VERSION : 0.1
   VAR
      VFD_DELAY : Array[1..5] of IEC_TIMER;
   END_VAR
BEGIN
   VFD_DELAY[1].PT := T#10S;
   VFD_DELAY[2].PT := T#10S;
END_DATA_BLOCK

// folder: Timers/Totalizer/Datablocks

DATA_BLOCK "FT-1045_Totalizer_DB"   // DB7
{ S7_Optimized_Access := 'TRUE' }
VERSION : 0.1
// stored: InstanceOfName Totalizer_1
"Totalizer_1"
BEGIN
   interval := T#30s;
   cycle := T#500ms;
END_DATA_BLOCK

DATA_BLOCK "FT-1041_Totalizer_DB"   // DB88
{ S7_Optimized_Access := 'TRUE' }
VERSION : 0.1
// stored: InstanceOfName Totalizer_1
"Totalizer_1"
BEGIN
   cycle := T#500ms;
   interval := T#30s;
END_DATA_BLOCK

DATA_BLOCK "FT-2022_Totalizer_DB"   // DB111
{ S7_Optimized_Access := 'TRUE' }
VERSION : 0.1
// stored: InstanceOfName Totalizer_1
"Totalizer_1"
BEGIN
   cycle := T#500ms;
   interval := T#30s;
END_DATA_BLOCK

DATA_BLOCK "FT-2012_Totalizer_DB"   // DB112
{ S7_Optimized_Access := 'TRUE' }
VERSION : 0.1
// stored: InstanceOfName Totalizer_1
"Totalizer_1"
BEGIN
   interval := T#30s;
   cycle := T#500ms;
END_DATA_BLOCK

DATA_BLOCK "FT-2011_Totalizer_DB"   // DB113
{ S7_Optimized_Access := 'TRUE' }
VERSION : 0.1
// stored: InstanceOfName Totalizer_1
"Totalizer_1"
BEGIN
   interval := T#30s;
   cycle := T#500ms;
END_DATA_BLOCK

DATA_BLOCK "FT-1044_Totalizer_DB"   // DB114
{ S7_Optimized_Access := 'TRUE' }
VERSION : 0.1
// stored: InstanceOfName Totalizer_1
"Totalizer_1"
BEGIN
   interval := T#30s;
   cycle := T#500ms;
END_DATA_BLOCK

DATA_BLOCK "FT-1043_Totalizer_DB"   // DB115
{ S7_Optimized_Access := 'TRUE' }
VERSION : 0.1
// stored: InstanceOfName Totalizer_1
"Totalizer_1"
BEGIN
   interval := T#30s;
   cycle := T#500ms;
END_DATA_BLOCK

DATA_BLOCK "FT-1042_Totalizer_DB"   // DB116
{ S7_Optimized_Access := 'TRUE' }
VERSION : 0.1
// stored: InstanceOfName Totalizer_1
"Totalizer_1"
BEGIN
   interval := T#30s;
   cycle := T#500ms;
END_DATA_BLOCK

DATA_BLOCK "FT-3011_Totalizer_DB"   // DB117
{ S7_Optimized_Access := 'TRUE' }
VERSION : 0.1
// stored: InstanceOfName Totalizer_1
"Totalizer_1"
BEGIN
   interval := T#30s;
   cycle := T#500MS;
END_DATA_BLOCK

DATA_BLOCK "FT-2021_Totalizer_DB"   // DB118
{ S7_Optimized_Access := 'TRUE' }
VERSION : 0.1
// stored: InstanceOfName Totalizer_1
"Totalizer_1"
BEGIN
   interval := T#30s;
   cycle := T#500ms;
END_DATA_BLOCK

DATA_BLOCK "FT-1021_Totalizer_DB"   // DB190
{ S7_Optimized_Access := 'TRUE' }
VERSION : 0.1
// stored: InstanceOfName Totalizer_1
"Totalizer_1"
BEGIN
   interval := T#30s;
   cycle := T#500ms;
END_DATA_BLOCK

DATA_BLOCK "FT-1011_Totalizer_DB"   // DB254
{ S7_Optimized_Access := 'TRUE' }
VERSION : 0.1
// stored: InstanceOfName Totalizer_1
"Totalizer_1"
BEGIN
END_DATA_BLOCK

DATA_BLOCK "FT-3012_Totalizer_DB"   // DB376
{ S7_Optimized_Access := 'TRUE' }
VERSION : 0.1
// stored: InstanceOfName Totalizer_1
"Totalizer_1"
BEGIN
   interval := T#30s;
   cycle := T#500ms;
END_DATA_BLOCK

// folder: VFD/Datablocks

DATA_BLOCK "VFD-C301_DB"   // DB1
{ S7_Optimized_Access := 'TRUE' }
VERSION : 0.7
// stored: InstanceOfName VFD_Dumbdown
"VFD_Dumbdown"
BEGIN
END_DATA_BLOCK

DATA_BLOCK "VFD-C301R_DB"   // DB84
{ S7_Optimized_Access := 'TRUE' }
VERSION : 0.7
// stored: InstanceOfName VFD_Dumbdown
"VFD_Dumbdown"
BEGIN
END_DATA_BLOCK

DATA_BLOCK "VFD-R201_DB"   // DB85
{ S7_Optimized_Access := 'TRUE' }
VERSION : 0.7
// stored: InstanceOfName VFD_Dumbdown
"VFD_Dumbdown"
BEGIN
   Motor_max_RPM := 450.0;
END_DATA_BLOCK

DATA_BLOCK "VFD-T103_DB"   // DB107
{ S7_Optimized_Access := 'TRUE' }
VERSION : 0.7
// stored: InstanceOfName VFD_Dumbdown
"VFD_Dumbdown"
BEGIN
END_DATA_BLOCK

DATA_BLOCK "VFD-T102A_DB"   // DB108
{ S7_Optimized_Access := 'TRUE' }
VERSION : 0.7
// stored: InstanceOfName VFD_Dumbdown
"VFD_Dumbdown"
BEGIN
   Motor_max_RPM := 1770.0;
END_DATA_BLOCK

DATA_BLOCK "VFD-T101A_DB"   // DB109
{ S7_Optimized_Access := 'TRUE' }
VERSION : 0.7
// stored: InstanceOfName VFD_Dumbdown
"VFD_Dumbdown"
BEGIN
   Motor_max_RPM := 1730.0;
END_DATA_BLOCK

DATA_BLOCK "VFD-R202_DB"   // DB110
{ S7_Optimized_Access := 'TRUE' }
VERSION : 0.7
// stored: InstanceOfName VFD_Dumbdown
"VFD_Dumbdown"
BEGIN
   Motor_max_RPM := 450.0;
END_DATA_BLOCK

DATA_BLOCK "VFD-T101B_DB"   // DB183
{ S7_Optimized_Access := 'TRUE' }
VERSION : 0.7
// stored: InstanceOfName VFD_Dumbdown
"VFD_Dumbdown"
BEGIN
   Motor_max_RPM := 1730.0;
END_DATA_BLOCK

DATA_BLOCK "VFD-T102B_DB"   // DB184
{ S7_Optimized_Access := 'TRUE' }
VERSION : 0.7
// stored: InstanceOfName VFD_Dumbdown
"VFD_Dumbdown"
BEGIN
   Motor_max_RPM := 1770.0;
END_DATA_BLOCK

// folder: VFD/T103_VFD

DATA_BLOCK "T103_VFD_Control_DB"   // DB263
{ S7_Optimized_Access := 'TRUE' }
VERSION : 0.1
   VAR
      AutoSpeedSP : Real;   // Auto Speed SP
   END_VAR
BEGIN
END_DATA_BLOCK

DATA_BLOCK "VFD_T103_PN_DB"   // DB264
{ S7_Optimized_Access := 'TRUE' }
VERSION : 0.1
// stored: InstanceOfName VFD_PNCtrl
"VFD_PNCtrl"
BEGIN
END_DATA_BLOCK

// folder: Valves/Control Valves

DATA_BLOCK "FV-4012_DB"   // DB177
{ S7_Optimized_Access := 'TRUE' }
VERSION : 0.1
// stored: InstanceOfName Valve-CV
"Valve-CV"
BEGIN
END_DATA_BLOCK

// folder: Valves/Control Valves/Datablocks

DATA_BLOCK "FV-2011_DB"   // DB80
{ S7_Optimized_Access := 'TRUE' }
VERSION : 0.1
// stored: InstanceOfName Valve-CV
"Valve-CV"
BEGIN
END_DATA_BLOCK

DATA_BLOCK "FV-2012_DB"   // DB81
{ S7_Optimized_Access := 'TRUE' }
VERSION : 0.1
// stored: InstanceOfName Valve-CV
"Valve-CV"
BEGIN
END_DATA_BLOCK

DATA_BLOCK "FV-2021_DB"   // DB82
{ S7_Optimized_Access := 'TRUE' }
VERSION : 0.1
// stored: InstanceOfName Valve-CV
"Valve-CV"
BEGIN
END_DATA_BLOCK

DATA_BLOCK "FV-2022_DB"   // DB83
{ S7_Optimized_Access := 'TRUE' }
VERSION : 0.1
// stored: InstanceOfName Valve-CV
"Valve-CV"
BEGIN
END_DATA_BLOCK

DATA_BLOCK "FV-3011_DB"   // DB234
{ S7_Optimized_Access := 'TRUE' }
VERSION : 0.1
// stored: InstanceOfName Valve-CV
"Valve-CV"
BEGIN
END_DATA_BLOCK

DATA_BLOCK "FV-4011_DB"   // DB381
{ S7_Optimized_Access := 'TRUE' }
VERSION : 0.1
// stored: InstanceOfName Valve-CV
"Valve-CV"
BEGIN
END_DATA_BLOCK

DATA_BLOCK "FV-4021_DB"   // DB418
{ S7_Optimized_Access := 'TRUE' }
VERSION : 0.1
// stored: InstanceOfName Valve-CV
"Valve-CV"
BEGIN
END_DATA_BLOCK

DATA_BLOCK "FV-4024_DB"   // DB419
{ S7_Optimized_Access := 'TRUE' }
VERSION : 0.1
// stored: InstanceOfName Valve-CV
"Valve-CV"
BEGIN
END_DATA_BLOCK

DATA_BLOCK "FV-4025_DB"   // DB420
{ S7_Optimized_Access := 'TRUE' }
VERSION : 0.1
// stored: InstanceOfName Valve-CV
"Valve-CV"
BEGIN
END_DATA_BLOCK

// folder: Valves/Solenoid Valve/Datablocks

DATA_BLOCK "XV-1033_DB"   // DB2
{ S7_Optimized_Access := 'FALSE' }
VERSION : 1.0
// stored: InstanceOfName Valve-SV
"Valve-SV"
BEGIN
   EM := 1;
END_DATA_BLOCK

DATA_BLOCK "XV-1041_DB"   // DB3
{ S7_Optimized_Access := 'FALSE' }
VERSION : 1.0
// stored: InstanceOfName Valve-SV
"Valve-SV"
BEGIN
   EM := 1;
END_DATA_BLOCK

DATA_BLOCK "XV-1011_DB"   // DB4
{ S7_Optimized_Access := 'FALSE' }
VERSION : 1.0
// stored: InstanceOfName Valve-SV
"Valve-SV"
BEGIN
   EM := 1;
END_DATA_BLOCK

DATA_BLOCK "XV-1013_DB"   // DB5
{ S7_Optimized_Access := 'FALSE' }
VERSION : 1.0
// stored: InstanceOfName Valve-SV
"Valve-SV"
BEGIN
   EM := 1;
END_DATA_BLOCK

DATA_BLOCK "XV-1021_DB"   // DB10
{ S7_Optimized_Access := 'FALSE' }
VERSION : 1.0
// stored: InstanceOfName Valve-SV
"Valve-SV"
BEGIN
   EM := 1;
END_DATA_BLOCK

DATA_BLOCK "XV-1043_DB"   // DB12
{ S7_Optimized_Access := 'FALSE' }
VERSION : 1.0
// stored: InstanceOfName Valve-SV
"Valve-SV"
BEGIN
   EM := 1;
END_DATA_BLOCK

DATA_BLOCK "XV-1044_DB"   // DB13
{ S7_Optimized_Access := 'FALSE' }
VERSION : 1.0
// stored: InstanceOfName Valve-SV
"Valve-SV"
BEGIN
   EM := 1;
END_DATA_BLOCK

DATA_BLOCK "XV-2011_DB"   // DB14
{ S7_Optimized_Access := 'FALSE' }
VERSION : 1.0
// stored: InstanceOfName Valve-SV
"Valve-SV"
BEGIN
   EM := 1;
END_DATA_BLOCK

DATA_BLOCK "XV-2012_DB"   // DB15
{ S7_Optimized_Access := 'FALSE' }
VERSION : 1.0
// stored: InstanceOfName Valve-SV
"Valve-SV"
BEGIN
   EM := 1;
END_DATA_BLOCK

DATA_BLOCK "XV-2013_DB"   // DB16
{ S7_Optimized_Access := 'FALSE' }
VERSION : 1.0
// stored: InstanceOfName Valve-SV
"Valve-SV"
BEGIN
   EM := 1;
END_DATA_BLOCK

DATA_BLOCK "XV-2021_DB"   // DB18
{ S7_Optimized_Access := 'FALSE' }
VERSION : 1.0
// stored: InstanceOfName Valve-SV
"Valve-SV"
BEGIN
   EM := 1;
END_DATA_BLOCK

DATA_BLOCK "XV-2023_DB"   // DB19
{ S7_Optimized_Access := 'FALSE' }
VERSION : 1.0
// stored: InstanceOfName Valve-SV
"Valve-SV"
BEGIN
   EM := 1;
END_DATA_BLOCK

DATA_BLOCK "XV-1032_DB"   // DB21
{ S7_Optimized_Access := 'FALSE' }
VERSION : 1.0
// stored: InstanceOfName Valve-SV
"Valve-SV"
BEGIN
   EM := 1;
END_DATA_BLOCK

DATA_BLOCK "XV-3011_DB"   // DB22
{ S7_Optimized_Access := 'FALSE' }
VERSION : 1.0
// stored: InstanceOfName Valve-SV
"Valve-SV"
BEGIN
   EM := 1;
END_DATA_BLOCK

DATA_BLOCK "XV-3012_DB"   // DB23
{ S7_Optimized_Access := 'FALSE' }
VERSION : 1.0
// stored: InstanceOfName Valve-SV
"Valve-SV"
BEGIN
   EM := 1;
END_DATA_BLOCK

DATA_BLOCK "XV-3013_DB"   // DB24
{ S7_Optimized_Access := 'FALSE' }
VERSION : 1.0
// stored: InstanceOfName Valve-SV
"Valve-SV"
BEGIN
   EM := 1;
END_DATA_BLOCK

DATA_BLOCK "XV-1045_DB"   // DB25
{ S7_Optimized_Access := 'FALSE' }
VERSION : 1.0
// stored: InstanceOfName Valve-SV
"Valve-SV"
BEGIN
   EM := 1;
END_DATA_BLOCK

DATA_BLOCK "XV-1023_DB"   // DB27
{ S7_Optimized_Access := 'FALSE' }
VERSION : 1.0
// stored: InstanceOfName Valve-SV
"Valve-SV"
BEGIN
   EM := 1;
END_DATA_BLOCK

DATA_BLOCK "XV-4024_DB"   // DB28
{ S7_Optimized_Access := 'FALSE' }
VERSION : 1.0
// stored: InstanceOfName Valve-SV
"Valve-SV"
BEGIN
   EM := 1;
END_DATA_BLOCK

DATA_BLOCK "XV-4025_DB"   // DB29
{ S7_Optimized_Access := 'FALSE' }
VERSION : 1.0
// stored: InstanceOfName Valve-SV
"Valve-SV"
BEGIN
   EM := 1;
END_DATA_BLOCK

DATA_BLOCK "XV-1042_DB"   // DB99
{ S7_Optimized_Access := 'FALSE' }
VERSION : 1.0
// stored: InstanceOfName Valve-SV
"Valve-SV"
BEGIN
   EM := 1;
END_DATA_BLOCK

DATA_BLOCK "XV-2022_DB"   // DB104
{ S7_Optimized_Access := 'FALSE' }
VERSION : 1.0
// stored: InstanceOfName Valve-SV
"Valve-SV"
BEGIN
   EM := 1;
END_DATA_BLOCK

DATA_BLOCK "XV-1031_DB"   // DB106
{ S7_Optimized_Access := 'FALSE' }
VERSION : 1.0
// stored: InstanceOfName Valve-SV
"Valve-SV"
BEGIN
   EM := 1;
END_DATA_BLOCK

DATA_BLOCK "XV-4021_DB"   // DB416
{ S7_Optimized_Access := 'FALSE' }
VERSION : 1.0
// stored: InstanceOfName Valve-SV
"Valve-SV"
BEGIN
END_DATA_BLOCK

DATA_BLOCK "XV-4022_DB"   // DB417
{ S7_Optimized_Access := 'FALSE' }
VERSION : 1.0
// stored: InstanceOfName Valve-SV
"Valve-SV"
BEGIN
END_DATA_BLOCK

// folder: 0)Organization Blocks

ORGANIZATION_BLOCK "Main"   // OB1, LAD, ProgramCycle
TITLE = "Main Program Sweep (Cycle)"
{ S7_Optimized_Access := 'TRUE' }
VERSION : 0.1
// Updated Date:
// Note:
   VAR_INPUT
      Initial_Call : Bool;   // Initial call of this OB
      Remanence : Bool;   // =True, if remanent data are available
   END_VAR
   VAR_TEMP
      "bool" : Bool;
   END_VAR
   VAR CONSTANT
      Idle_Star : Int := 0;
      Idle_End : Int := 49;
      Shutdown_Star : Int := 50;
      Shutdown_End : Int := 99;
      Inititilize_Start : Int := 100;
      Inititilize_End : Int := 199;
   END_VAR
BEGIN

REGION Network 1: Interlocks & Diagnostic
   // Interlocks_FC: Contains all interlock Sequences 
   // Diag_FC: Contains all diagnostic  Sequences
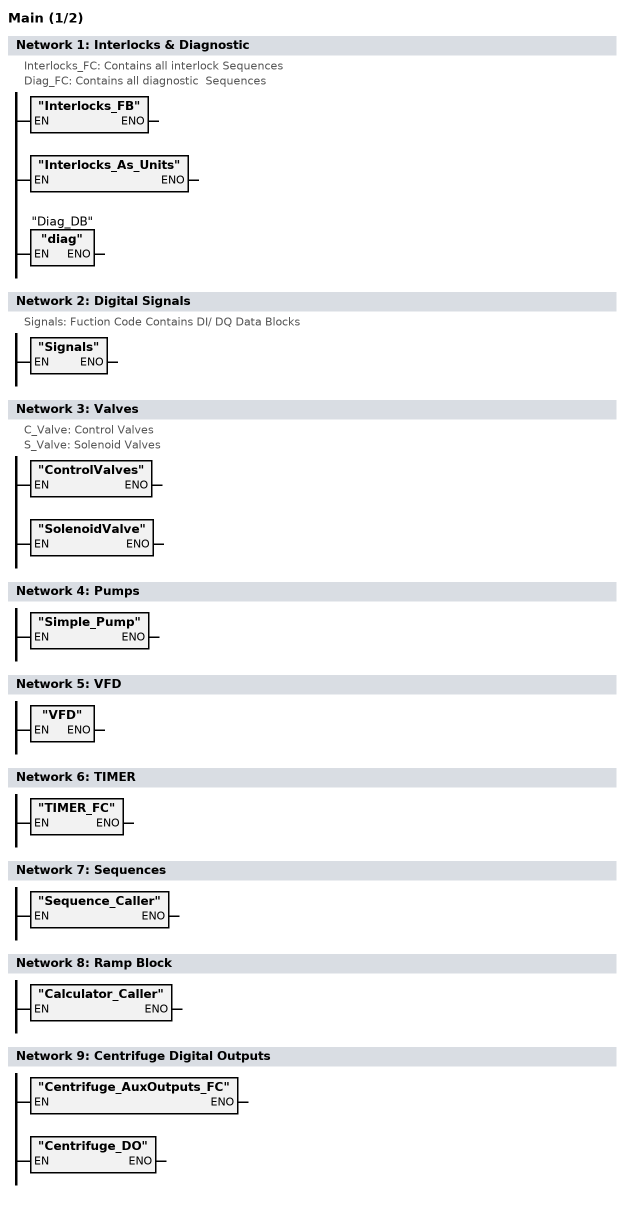
   RUNG wire#powerrail
      "Interlocks_FB"()
   END_RUNG
   RUNG wire#powerrail
      "Interlocks_As_Units"()
   END_RUNG
   RUNG wire#powerrail
      "Diag_DB"()
   END_RUNG
   // the same network as SCL:
   "Interlocks_FB"();
   "Interlocks_As_Units"();
   "Diag_DB"();   // "diag"
END_REGION

REGION Network 2: Digital Signals
   // Signals: Fuction Code Contains DI/ DQ Data Blocks
   RUNG wire#powerrail
      "Signals"()
   END_RUNG
   // the same network as SCL:
   "Signals"();
END_REGION

REGION Network 3: Valves
   // C_Valve: Control Valves 
   // S_Valve: Solenoid Valves
   RUNG wire#powerrail
      "ControlValves"()
   END_RUNG
   RUNG wire#powerrail
      "SolenoidValve"()
   END_RUNG
   // the same network as SCL:
   "ControlValves"();
   "SolenoidValve"();
END_REGION

REGION Network 4: Pumps
   RUNG wire#powerrail
      "Simple_Pump"()
   END_RUNG
   // the same network as SCL:
   "Simple_Pump"();
END_REGION

REGION Network 5: VFD
   RUNG wire#powerrail
      "VFD"()
   END_RUNG
   // the same network as SCL:
   "VFD"();
END_REGION

REGION Network 6: TIMER
   RUNG wire#powerrail
      "TIMER_FC"()
   END_RUNG
   // the same network as SCL:
   "TIMER_FC"();
END_REGION

REGION Network 7: Sequences
   RUNG wire#powerrail
      "Sequence_Caller"()
   END_RUNG
   // the same network as SCL:
   "Sequence_Caller"();
END_REGION

REGION Network 8: Ramp Block
   RUNG wire#powerrail
      "Calculator_Caller"()
   END_RUNG
   // the same network as SCL:
   "Calculator_Caller"();
END_REGION

REGION Network 9: Centrifuge Digital Outputs
   RUNG wire#powerrail
      "Centrifuge_AuxOutputs_FC"()
   END_RUNG
   RUNG wire#powerrail
      "Centrifuge_DO"()
   END_RUNG
   // the same network as SCL:
   "Centrifuge_AuxOutputs_FC"();
   "Centrifuge_DO"();
END_REGION

REGION Network 10: Cause and Effect Matrix
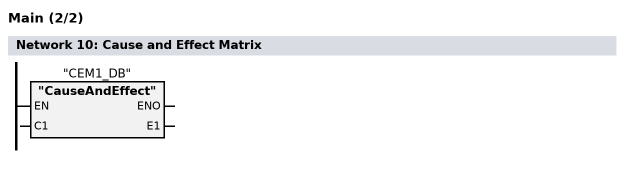
   RUNG wire#powerrail
      "CEM1_DB"(C1 :=, E1 =>)
   END_RUNG
   // the same network as SCL:
   "CEM1_DB"();   // "CauseAndEffect"
END_REGION
END_ORGANIZATION_BLOCK

ORGANIZATION_BLOCK "Cycle_5s"   // OB30, LAD, CyclicInterrupt
{ S7_Optimized_Access := 'TRUE' }
VERSION : 0.1
   VAR_INPUT
      Initial_Call : Bool;   // Initial call of this OB
      Event_Count : Int;   // Events discarded
   END_VAR
BEGIN

REGION Network 1: Temperature Trasmitters
   // Temperature Trasmitters Function Code
END_REGION
END_ORGANIZATION_BLOCK

ORGANIZATION_BLOCK "Cycle_100ms"   // OB31, LAD, CyclicInterrupt
{ S7_Optimized_Access := 'TRUE' }
VERSION : 0.1
   VAR_INPUT
      Initial_Call : Bool;   // Initial call of this OB
      Event_Count : Int;   // Events discarded
   END_VAR
   VAR_TEMP   // added for the SCL form of the ladder/FBD networks
      _w1 : Bool;
      _w2 : Bool;
      _w3 : Bool;
   END_VAR
BEGIN

REGION Network 1: PH Trasmitters
   // PH Trasmitters Function Code
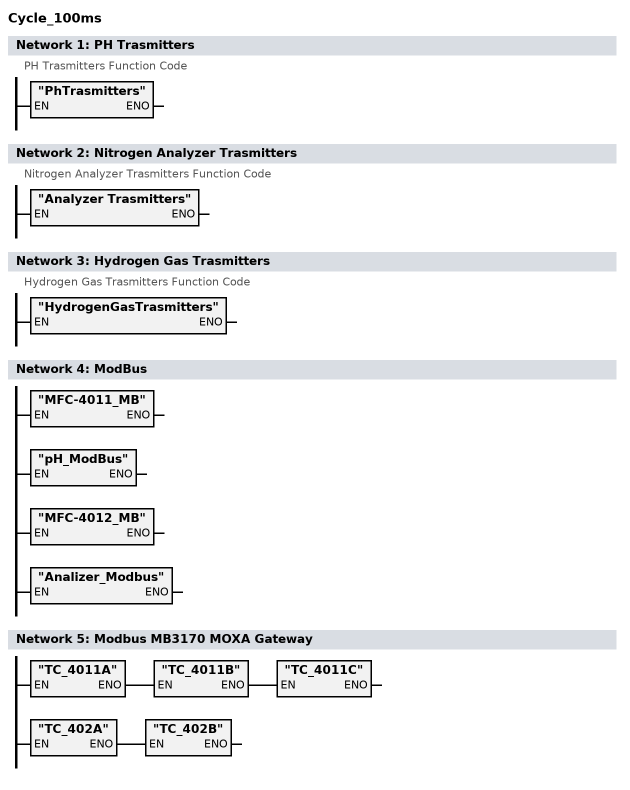
   RUNG wire#powerrail
      "PhTrasmitters"()
   END_RUNG
   // the same network as SCL:
   "PhTrasmitters"();
END_REGION

REGION Network 2: Nitrogen Analyzer Trasmitters
   // Nitrogen Analyzer Trasmitters Function Code
   RUNG wire#powerrail
      "Analyzer Trasmitters"()
   END_RUNG
   // the same network as SCL:
   "Analyzer Trasmitters"();
END_REGION

REGION Network 3: Hydrogen Gas Trasmitters
   // Hydrogen Gas Trasmitters Function Code
   RUNG wire#powerrail
      "HydrogenGasTrasmitters"()
   END_RUNG
   // the same network as SCL:
   "HydrogenGasTrasmitters"();
END_REGION

REGION Network 4: ModBus
   RUNG wire#powerrail
      "MFC-4011_MB"()
   END_RUNG
   RUNG wire#powerrail
      "pH_ModBus"()
   END_RUNG
   RUNG wire#powerrail
      "MFC-4012_MB"()
   END_RUNG
   RUNG wire#powerrail
      "Analizer_Modbus"()
   END_RUNG
   // the same network as SCL:
   "MFC-4011_MB"();
   "pH_ModBus"();
   "MFC-4012_MB"();
   "Analizer_Modbus"();
END_REGION

REGION Network 5: Modbus MB3170 MOXA Gateway
   RUNG wire#powerrail
      "TC_4011A"()
      "TC_4011B"()
      "TC_4011C"()
   END_RUNG
   RUNG wire#powerrail
      "TC_402A"()
      "TC_402B"()
   END_RUNG
   // the same network as SCL:
   "TC_4011A"(ENO => #_w1);
   "TC_4011B"(EN := #_w1, ENO => #_w2);
   IF #_w2 THEN "TC_4011C"(); END_IF;
   "TC_402A"(ENO => #_w3);
   IF #_w3 THEN "TC_402B"(); END_IF;
END_REGION
END_ORGANIZATION_BLOCK

ORGANIZATION_BLOCK "Cycle_1s"   // OB32, LAD, CyclicInterrupt
TITLE = Cyclic interrupt (Cycle) 1 Second"
{ S7_Optimized_Access := 'TRUE' }
VERSION : 0.1
   VAR_INPUT
      Initial_Call : Bool;   // Initial call of this OB
      Event_Count : Int;   // Events discarded
   END_VAR
BEGIN

REGION Network 1: PIDController
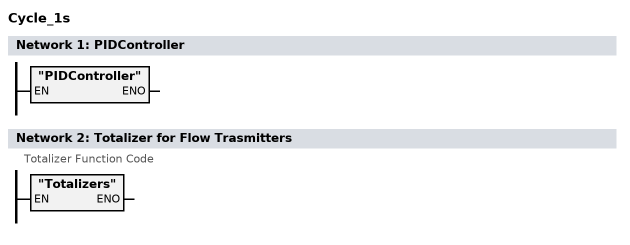
   RUNG wire#powerrail
      "PIDController"()
   END_RUNG
   // the same network as SCL:
   "PIDController"();
END_REGION

REGION Network 2: Totalizer for Flow Trasmitters
   // Totalizer Function Code
   RUNG wire#powerrail
      "Totalizers"()
   END_RUNG
   // the same network as SCL:
   "Totalizers"();
END_REGION
END_ORGANIZATION_BLOCK

ORGANIZATION_BLOCK "Cycle_500ms"   // OB33, LAD, CyclicInterrupt
{ S7_Optimized_Access := 'TRUE' }
VERSION : 0.1
   VAR_INPUT
      Initial_Call : Bool;   // Initial call of this OB
      Event_Count : Int;   // Events discarded
   END_VAR
   VAR_TEMP
      "REAL_R-201" : Real;
      "INT_R-201" : Real;
      "INT_R-202" : Real;
      "REAL_R-202" : Real;
   END_VAR
BEGIN

REGION Network 1: Flow Trasmitters
   // Flow Trasmitters Function Code
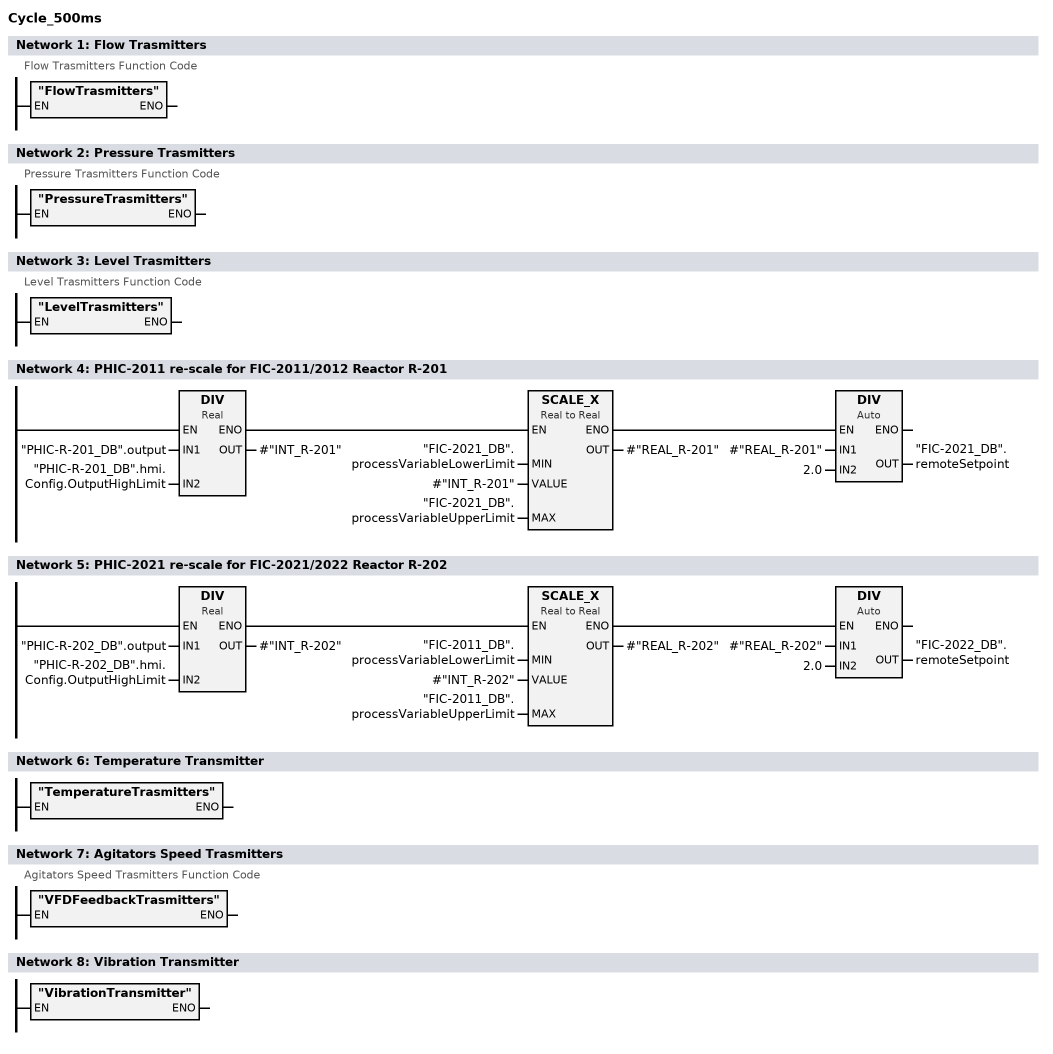
   RUNG wire#powerrail
      "FlowTrasmitters"()
   END_RUNG
   // the same network as SCL:
   "FlowTrasmitters"();
END_REGION

REGION Network 2: Pressure Trasmitters
   // Pressure Trasmitters Function Code
   RUNG wire#powerrail
      "PressureTrasmitters"()
   END_RUNG
   // the same network as SCL:
   "PressureTrasmitters"();
END_REGION

REGION Network 3: Level Trasmitters
   // Level Trasmitters Function Code
   RUNG wire#powerrail
      "LevelTrasmitters"()
   END_RUNG
   // the same network as SCL:
   "LevelTrasmitters"();
END_REGION

REGION Network 4: PHIC-2011 re-scale for FIC-2011/2012 Reactor R-201
   RUNG wire#powerrail
      { S7_Templates := "SrcType := Real"; S7_GenerateENO := "TRUE" } Div(in1 := "PHIC-R-201_DB".output, in2 := "PHIC-R-201_DB".hmi.Config.OutputHighLimit, out => #"INT_R-201")
      { S7_Templates := "[SrcType := Real, DestType := Real]"; S7_GenerateENO := "TRUE" } Scale(min := "FIC-2021_DB".processVariableLowerLimit, value := #"INT_R-201", max := "FIC-2021_DB".processVariableUpperLimit, out => #"REAL_R-201")
      { S7_GenerateENO := "TRUE" } Div(in1 := #"REAL_R-201", in2 := 2.0, out => "FIC-2021_DB".remoteSetpoint)
   END_RUNG
   // the same network as SCL:
   // ENO of a box is taken as its EN; it also drops when the box reports an error
   #"INT_R-201" := "PHIC-R-201_DB".output / "PHIC-R-201_DB".hmi.Config.OutputHighLimit;
   #"REAL_R-201" := SCALE_X(MIN := "FIC-2021_DB".processVariableLowerLimit, VALUE := #"INT_R-201", MAX := "FIC-2021_DB".processVariableUpperLimit);
   "FIC-2021_DB".remoteSetpoint := #"REAL_R-201" / 2.0;
END_REGION

REGION Network 5: PHIC-2021 re-scale for FIC-2021/2022 Reactor R-202
   RUNG wire#powerrail
      { S7_Templates := "SrcType := Real"; S7_GenerateENO := "TRUE" } Div(in1 := "PHIC-R-202_DB".output, in2 := "PHIC-R-202_DB".hmi.Config.OutputHighLimit, out => #"INT_R-202")
      { S7_Templates := "[SrcType := Real, DestType := Real]"; S7_GenerateENO := "TRUE" } Scale(min := "FIC-2011_DB".processVariableLowerLimit, value := #"INT_R-202", max := "FIC-2011_DB".processVariableUpperLimit, out => #"REAL_R-202")
      { S7_GenerateENO := "TRUE" } Div(in1 := #"REAL_R-202", in2 := 2.0, out => "FIC-2022_DB".remoteSetpoint)
   END_RUNG
   // the same network as SCL:
   // ENO of a box is taken as its EN; it also drops when the box reports an error
   #"INT_R-202" := "PHIC-R-202_DB".output / "PHIC-R-202_DB".hmi.Config.OutputHighLimit;
   #"REAL_R-202" := SCALE_X(MIN := "FIC-2011_DB".processVariableLowerLimit, VALUE := #"INT_R-202", MAX := "FIC-2011_DB".processVariableUpperLimit);
   "FIC-2022_DB".remoteSetpoint := #"REAL_R-202" / 2.0;
END_REGION

REGION Network 6: Temperature Transmitter
   RUNG wire#powerrail
      "TemperatureTrasmitters"()
   END_RUNG
   // the same network as SCL:
   "TemperatureTrasmitters"();
END_REGION

REGION Network 7: Agitators Speed Trasmitters
   // Agitators Speed Trasmitters Function Code
   RUNG wire#powerrail
      "VFDFeedbackTrasmitters"()
   END_RUNG
   // the same network as SCL:
   "VFDFeedbackTrasmitters"();
END_REGION

REGION Network 8: Vibration Transmitter
   RUNG wire#powerrail
      "VibrationTransmitter"()
   END_RUNG
   // the same network as SCL:
   "VibrationTransmitter"();
END_REGION
END_ORGANIZATION_BLOCK

ORGANIZATION_BLOCK "CPU redundancy error"   // OB72, LAD, CPURedundancyError
{ S7_Optimized_Access := 'TRUE' }
VERSION : 0.1
   VAR_INPUT
      LADDR : Hw_Any;   // Hardware identifier of the local device
      Event_Class : Byte;   // according to S7 classic
      Fault_ID : Byte;   // Fault_ID as in S7 classic
   END_VAR
BEGIN
END_ORGANIZATION_BLOCK

ORGANIZATION_BLOCK "Diagnostic error interrupt"   // OB82, LAD, DiagnosticErrorInterrupt
{ S7_Optimized_Access := 'TRUE' }
VERSION : 0.1
   VAR_INPUT
      IO_State : Word;   // IO state of the HW object
      LADDR : Hw_Any;   // Hardware identifier
      Channel : UInt;   // Channel number
      MultiError : Bool;   // =true if more than one error is present
   END_VAR
BEGIN
END_ORGANIZATION_BLOCK

ORGANIZATION_BLOCK "Startup"   // OB100, LAD, Startup
TITLE = "Complete Restart"
{ S7_Optimized_Access := 'TRUE' }
VERSION : 0.1
   VAR_INPUT
      LostRetentive : Bool;   // True if retentive data are lost
      LostRTC : Bool;   // True if date and time are lost
   END_VAR
BEGIN

REGION Network 1: VFD Set to Automode
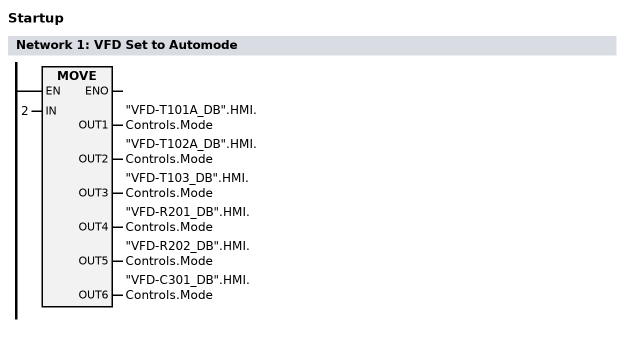
   RUNG wire#powerrail
      { S7_GenerateENO := "TRUE" } Move(in := 2, out1 => "VFD-T101A_DB".HMI.Controls.Mode, out2 => "VFD-T102A_DB".HMI.Controls.Mode, out3 => "VFD-T103_DB".HMI.Controls.Mode, out4 => "VFD-R201_DB".HMI.Controls.Mode, out5 => "VFD-R202_DB".HMI.Controls.Mode, out6 => "VFD-C301_DB".HMI.Controls.Mode)
   END_RUNG
   // the same network as SCL:
   "VFD-T101A_DB".HMI.Controls.Mode := 2;
   "VFD-T102A_DB".HMI.Controls.Mode := 2;
   "VFD-T103_DB".HMI.Controls.Mode := 2;
   "VFD-R201_DB".HMI.Controls.Mode := 2;
   "VFD-R202_DB".HMI.Controls.Mode := 2;
   "VFD-C301_DB".HMI.Controls.Mode := 2;
END_REGION
END_ORGANIZATION_BLOCK

ORGANIZATION_BLOCK "Programming error"   // OB121, LAD, ProgrammingError
{ S7_Optimized_Access := 'TRUE' }
VERSION : 0.1
   VAR_INPUT
      BlockNr : UInt;   // Number of causing block
      Reaction : USInt;   // 0:ignore, 1:substitute, 2:skip
      Fault_ID : Byte;   // Fault identifier
      BlockType : USInt;   // 16#01:OB, 16#02:FC, 16#03:FB, 16#04:SFC, 16#05:SFB, 16#06:DB: Type of block causing the error
      Area : USInt;   // Area where the error occured
      DBNr : DB_ANY;   // DB number if Area = DB or DI
      Csg_OBNr : OB_Any;   // Number of OB causing the error
      Csg_Prio : USInt;   // Priority of OB causing the error
      Width : USInt;   // 0:bit, 1:byte, 2:word, 3:dword, 4:lword
   END_VAR
BEGIN
END_ORGANIZATION_BLOCK

ORGANIZATION_BLOCK "IO access error"   // OB122, LAD, IOAccessError
{ S7_Optimized_Access := 'TRUE' }
VERSION : 0.1
   VAR_INPUT
      BlockNr : UInt;   // Number of causing block
      Reaction : USInt;   // 0:ignore, 1:substitute, 2:skip
      Fault_ID : Byte;   // 16#42:reading, 16#43:writing
      BlockType : USInt;   // 16#01:OB, 16#02:FC, 16#03:FB, 16#04:SFC, 16#05:SFB, 16#06:DB: Type of block causing the error
      Area : USInt;   // 16#81:I, 16#82:Q: IO area where the IOaccess error occured
      DBNr : DB_ANY;   // Reserved for system
      Csg_OBNr : OB_Any;   // Number of OB causing the error
      Csg_Prio : USInt;   // Priority of OB causing the error
      Width : USInt;   // 0:bit, 1:byte, 2:word, 3:dword, 4:lword
   END_VAR
BEGIN
END_ORGANIZATION_BLOCK

// folder: 1}Library

FUNCTION_BLOCK "UPS1600"   // FB15, LAD
{ S7_Optimized_Access := 'TRUE' }
VERSION : 0.1
   VAR_INPUT
      addrIn : Hw_Io := 260;   // HW-address of the UPS1600 must be insert there
      cyclicIOAddr : Hw_Io;   // IO Data submodule address must be inserted here
      upsExecuteReset : Bool;   // Input must be set if the station is ready for shutdown <- the station/ partners are ready to deactivate the tension
   END_VAR
   VAR_OUTPUT
      upsReadyForReset : Bool := False;   // Output will be set if the Block timer elapse -> signal to shutdown the station/ partners
   END_VAR
   VAR
      HMI : Struct
         Mode : Struct
            bufferMode : Byte := 16#80;   // Buffer mode //Value range: 0 = active, 255 = inactive
            readyForBuffering : Byte;   // Buffer readiness //Value range: 0=FALSE, 255=TRUE
         END_STRUCT;
         State : Struct
            Details : Struct
               orderNumber : String[20];   // Article no.
               serialNumber : String[20];   // Serial number
               deviceName : String[20];   // Name of the device
               versionNumber : String[30];   // Version number
               deviceHwRevision : Int;   // HW revision
               deviceSwRevision1 : Byte;   // SW revision1
               deviceSwRevision2 : Byte;   // SW revision2
               deviceSwRevision3 : Byte;   // Sw revision3
               batFamily : Byte;   // Battery family //Value range: BAT1600 = 1, UPS1100 = 2, Third-party battery = 3
               commandID : Int;   // Remote reset : 8207
               parameter1 : Byte;   // Waiting time after end of communication [s]
               parameter2 : Byte;   // output voltage down time [s]
            END_STRUCT;
            numOfBatteries : Byte;   // Number of batteries //Value range: 0 -6
            batteryType : Byte;   // Type of battery identifier //Value range: Pb =0, Li = 1
            inputVolt : Real;   // Input voltage //Value range: [0.01V]
            inputCur : Real;   // Input current //Value range: [5mA]
            outputVolt : Real;   // Output voltage //Value range: [0.01V]
            outputCur : Real;   // Output current //Value range: [5mA]
            maxOutCur : Byte;   // Maximum output current //Value range: [mA]
            bufferTime : Int;   // Buffer time //Value range: 1 - 32767s
            bufferThreshold : Real;   // Connection threshold //Value range: 21 - 25V
            bufferingAllowed : Byte;   // Buffering allowed //Value range: 0=FALSE, 255=TRUE
            batteryVolt : Real;   // Battery voltage //Value range: [0.01V]
            batteryChargeLevel : Byte := B#16#00;   // Battery charge level //Value range: 0 - 100%, 255 - unknown battery
            measuredChargeCur : Real;   // Measured charge current //Value range: [1mA]
            endOfChargeVolt : Real;   // End of charge voltage //Value range: 24 - 30V
            chargingOpState : Byte;   // Status of charging unit //Value range: 0 -4
            chargeVolt : Real;   // Current charge voltage //Value range: [0.01V]
            batteryDetails : Array[0..5] of Struct
               batteryLEDState : Byte;   // Signaling //Value range: Bit0/1: Color 0 = green/read alternating 1 = red 2 = green 3 = yellow Bit2/3: State 0 = off 1 = On 2 = 0,5Hz blinking 3 = 2Hz blinking
               batteryOpState : Byte;   // Battery status //Value range: 0 -11
               batteryCalcHealth : Byte;   // Calculated battery health //Value range: 0 -100
            END_STRUCT;
            totCalcBatCap : Real := 70.0;   // Calculated battery capacity [ 0.1Ah]
            loadCur : Real;   // Load current //Value range: [5mA]
         END_STRUCT;
      END_STRUCT;
      statBufferTime : Time := T#10S;   // time for the timer (default: 10s)
      statSetTimer : Bool;
      statBlockTimer : Bool;
      statDataBufParam : Struct   // Buffering Parameters
         bufferTime : Int := 600;   // Buffer time [s], AllowedValues = 1..32767
         bufferTime2 : Int := 60;   // Buffer time 2 [s], AllowedValues = 1..300
         bufferThreshold : Int := 2250;   // Buffer Threshold [0.01V], AllowedValues = 2100..2500
         stopBuffVoltage : Int := 1850;   // Stop Buffering Voltage [0.01V], AllowedValues = 1800..2300
         InputVoltOkTime : Int := 1000;   // Input Voltage OK Time [ms], AllowedValues = 200..65000
         downtimeAlarm : Int := 100;   // Downtime alarm [ms], AllowedValues = 0..20000
         bufferingAllowed : Byte := 16#FF;   // Buffering Allowed, AllowedValues = [0/255]
         enableResetAfterBuff : Byte := 16#00;   // Enable Reset after buffering , AllowedValues = [0/255]
         dischargeCutOffVolt : Int;
      END_STRUCT;
      statDataDeviceInfo : Struct   // Device Information
         hwRevision : Int;   // HW revision
         swRevision : Int;   // SW revision
         bootLoaderVersion : Int;   // Boot loader version
         maxOutCur : Byte;   // Maximum output current [A]
         padding : Byte;
         orderNumber : Array[0..18] of Char;   // MLFB/Order number
         serialNumber : Array[0..14] of Char;   // Serial number
         deviceName : Array[0..29] of Char;   // Device name
         versionNumber : Array[0..49] of Char;   // Version number
      END_STRUCT;
      statDataStateInfo : Struct   // State Information
         remainingBufferTime : DInt;   // Remaining buffer time [s]
         totalOperatingTime : DInt;   // Total operating time [hours]
         totalCalcBatCapacity : Int;   // Total calculated battery capacity [0.1Ah]
         calcBatCapacity : Array[0..5] of Int;   // Calculated battery capacity (battery 1 to 6) [0.1Ah]
         inputVolt : Int;   // Input voltage [0.01V]
         inputCur : Int;   // Input current [5mA]
         outputVolt : Int;   // Output voltage [0.01V]
         loadCur : Int;   // Load current [5mA]
         measuredChargeCur : Int;   // Measured charge current [mA]
         batteryVolt : Int;   // Battery voltage [0.01V]
         outputCur : Int;   // Output current [5mA]
         chargeVolt : Int;   // Charge voltage [0.01V]
         padding1 : Byte;
         padding2 : Byte;
         padding3 : Byte;
         validConfig : Byte;   // Valid configuration
         numOfBatteries : Byte;   // Number of batteries
         Reserved1 : Byte;
         Reserved2 : Byte;
         Reserved3 : Byte;
         Reserved4 : Byte;
         Reserved5 : Byte;
         Reserved6 : Byte;
         Reserved7 : Byte;
         bat1ChangeRecomm : Byte;   // Battery 1 change recommended
         bat2ChangeRecomm : Byte;   // Battery 2 change recommended
         bat3ChangeRecomm : Byte;   // Battery 3 change recommended
         bat4ChangeRecomm : Byte;   // Battery 4 change recommended
         bat5ChangeRecomm : Byte;   // Battery 5 change recommended
         bat6ChangeRecomm : Byte;   // Battery 6 change recommended
         bat1ConnFault : Byte;   // Battery 1 connection fault
         bat2ConnFault : Byte;   // Battery 2 connection fault
         bat3ConnFault : Byte;   // Battery 3 connection fault
         bat4ConnFault : Byte;   // Battery 4 connection fault
         bat5ConnFault : Byte;   // Battery 5 connection fault
         bat6ConnFault : Byte;   // Battery 6 connection fault
         bat1Temp : Byte;   // Battery 1 Temperature [1°C]
         bat2Temp : Byte;   // Battery 2 Temperature [1°C]
         bat3Temp : Byte;   // Battery 3 Temperature [1°C]
         bat4Temp : Byte;   // Battery 4 Temperature [1°C]
         bat5Temp : Byte;   // Battery 5 Temperature [1°C]
         bat6Temp : Byte;   // Battery 6 Temperature [1°C]
         deviceTemp : Byte;   // Device temperature [1°C]
         LEDPattern : Byte;   // LED pattern
         batCalBatHealth : Array[0..5] of Byte;
         batOpState : Array[0..5] of Byte;
         batLEDstate : Array[0..5] of Byte;
         chargingOpState : Byte;
      END_STRUCT;
      statDataUPSIandM : Struct   // I & M0 Handler
         blockHeader : Array[1..3] of Int;   // Block header
         vendorID : Int;   // Vendor ID
         orderId : Array[1..20] of Char;   // Order ID
         serNum : Array[1..16] of Char;   // Serial number
         hwRevision : Int;   // Device Product state
         swRevision : DWord;   // SW version of device
         revCnt : Int;   // RevCnt
         profId : Int;   // ProfID
         profSpecTyp : Int;   // ProfSpecTyp
         versMaj : Byte;   // VersMaj
         versMin : Byte;   // VersMin
         supported : Int;   // Supported
      END_STRUCT;
      statDataUPSCmd : Struct   // DC UPS Command
         commandID : Int := 8207;   // Remote reset2 = 8207 ; Output ON/OFF = 8200
         parameter1 : Byte := 16#3C;   // Buffer Time2 [s], AllowedValues = 1..300
         parameter2 : Byte := 16#05;   // Reset Time [s], AllowedValues = 1..120
      END_STRUCT;
      statDataResetParam : Byte := 16#05;   // Reset Time, AllowedValues = 1..120
      statRdReq : Bool;
      statWrReq : Bool;
      statValue : Int;
      statDataRecordRead : RDREC;
      statDataRecordBatInfo : RDREC;
      statDataRecordWrite : WRREC;
      statOrderNumberStr : String;   // Order number (String)
      statSerialNumberStr : String;   // Serial number (String)
      statDeviceNameStr : String;   // Device name (String)
      statVersionNumberStr : String;   // Version number (String)
      statCyclicData : Array[0..7] of Byte;
      statRetVal : DInt;
      statTimerObj : TON_TIME;
      statDataBatteryInfo : Struct
         numOfBatteries : Byte;
         padding1 : Byte;
         padding2 : Byte;
         padding3 : Byte;
         batteryDetails : Array[0..5] of Struct
            standbyTime : DInt;
            bufferTime : DInt;
            totChargingCur : DInt;
            totCulledCur : DInt;
            eocv : Int;
            chargeCur : Int;
            batCapacity : Int;
            stopBufVolt : Int;
            batteryType : Byte;
            minimalTemp : Byte;
            maximalTemp : Byte;
            orderNum : Array[0..18] of Char;
            serialNum : Array[0..14] of Char;
            manufacturingDate : Array[0..7] of Char;
            versionNum : Array[0..5] of Char;
            batCalcHealth : Byte;
            batOpState : Byte;
            batLEDState : Byte;
            padding4 : Byte;
            padding5 : Byte;
            batSWD : DWord;
            batMID : DWord;
         END_STRUCT;
      END_STRUCT;
      statStatusFLag1 : Byte;
      statStatusFLag2 : Byte;
      statCmdDone : Bool;   // 1 = Command writing is done, 0 = Command is not writtent to UPS1600
      statDevInfoRead : Byte;   // 1 = Device Info read, 0 = Device Info not read
      statBatteryFamily1 : Byte;
      statBatteryFamily2 : Byte;
      statCyclicCount : Int;
   END_VAR
   VAR_TEMP
      tempIterator : Int;
   END_VAR
   // // HMI.State.batteryDetails[1].batteryLEDState : Signaling //Value range: Bit0/1: Color 0 = green/read alternating 1 = red 2 = green 3 = yellow Bit2/3: State 0 = off 1 = On 2 = 0,5Hz blinking 3 = 2Hz blinking
   // // HMI.State.batteryDetails[2].batteryLEDState : Signaling //Value range: Bit0/1: Color 0 = green/read alternating 1 = red 2 = green 3 = yellow Bit2/3: State 0 = off 1 = On 2 = 0,5Hz blinking 3 = 2Hz blinking
   // // HMI.State.batteryDetails[3].batteryLEDState : Signaling //Value range: Bit0/1: Color 0 = green/read alternating 1 = red 2 = green 3 = yellow Bit2/3: State 0 = off 1 = On 2 = 0,5Hz blinking 3 = 2Hz blinking
   // // HMI.State.batteryDetails[4].batteryLEDState : Signaling //Value range: Bit0/1: Color 0 = green/read alternating 1 = red 2 = green 3 = yellow Bit2/3: State 0 = off 1 = On 2 = 0,5Hz blinking 3 = 2Hz blinking
   // // HMI.State.batteryDetails[5].batteryLEDState : Signaling //Value range: Bit0/1: Color 0 = green/read alternating 1 = red 2 = green 3 = yellow Bit2/3: State 0 = off 1 = On 2 = 0,5Hz blinking 3 = 2Hz blinking
   // // HMI.State.batteryDetails[1].batteryOpState : Battery status //Value range: 0 -11
   // // HMI.State.batteryDetails[2].batteryOpState : Battery status //Value range: 0 -11
   // // HMI.State.batteryDetails[3].batteryOpState : Battery status //Value range: 0 -11
   // // HMI.State.batteryDetails[4].batteryOpState : Battery status //Value range: 0 -11
   // // HMI.State.batteryDetails[5].batteryOpState : Battery status //Value range: 0 -11
   // // HMI.State.batteryDetails[1].batteryCalcHealth : Calculated battery health //Value range: 0 -100
   // // HMI.State.batteryDetails[2].batteryCalcHealth : Calculated battery health //Value range: 0 -100
   // // HMI.State.batteryDetails[3].batteryCalcHealth : Calculated battery health //Value range: 0 -100
   // // HMI.State.batteryDetails[4].batteryCalcHealth : Calculated battery health //Value range: 0 -100
   // // HMI.State.batteryDetails[5].batteryCalcHealth : Calculated battery health //Value range: 0 -100
BEGIN

REGION Network 1 (SCL): UPS1600 SCL Code
   //============================================================================= 
   // Copyright (C) Siemens AG 2020. All Rights Reserved. Confidential
   //----------------------------------------------------------------------------- 
   //Function block UPS1600 
   // Requirements: (hardware, technological package, memory needed, etc.) 
   // The functionality of the UPS1600 block is 
   //  - Reading Cyclic data records
   //  - Reading of acyclic data records
   //  - Writing of acyclic data records
   //  - Monitoring Buffer mode of UPS1600 and shutdown plant safely.
   //  

   //============================================================================= 
   //sequence chain (#statValue)
   // DW   2022-02-10  Moved the data structure from a udt to the static area and organized it more like the OA data structure.

   IF (#addrIn <> 0) AND (#cyclicIOAddr <> 0) THEN
       IF #statValue = 0 OR #statValue > 7 THEN
           #statValue := 1;
       END_IF;

       //cases of #statValue
       CASE #statValue OF
           1:
               IF NOT #statRdReq AND NOT #statDataRecordRead.BUSY THEN
                   #statRdReq := 1;
               END_IF;
               #statDataRecordRead(REQ := #statRdReq,  // IN: BOOL
                                   ID := #addrIn,  // IN: DINT
                                   INDEX := 32,  // IN: INT
                                   MLEN := 89, // IN: INT
                                   RECORD := #statDataStateInfo);  // INOUT: ANY

               IF NOT #statDataRecordRead.ERROR AND NOT #statDataRecordRead.BUSY THEN
                   IF #statStatusFLag1 < 1 THEN
                       #statStatusFLag1 := 1;
                   END_IF;
               END_IF;

               IF NOT #statDataRecordRead.BUSY OR #statDataRecordRead.ERROR THEN
                   #statRdReq := 0;
                   #statValue := 2;
               END_IF;

           2:
               IF NOT #statRdReq AND NOT #statDataRecordRead.BUSY THEN
                   #statRdReq := 1;
               END_IF;
               #statDataRecordRead(REQ := #statRdReq, // IN: BOOL
                                   ID := #addrIn,  // IN: DINT
                                   INDEX := 1,  // IN: INT
                                   MLEN := 16, // IN: INT
                                   RECORD := #statDataBufParam);  // INOUT: ANY

               IF NOT #statDataRecordRead.BUSY OR #statDataRecordRead.ERROR THEN
                   #statRdReq := 0;
                   #statValue := 3;
                   //END_IF;
               END_IF;

           3:
               IF NOT #statRdReq AND NOT #statDataRecordRead.BUSY THEN
                   #statRdReq := 1;
               END_IF;
               #statDataRecordRead(REQ := #statRdReq,  // IN: BOOL
                                   ID := #addrIn,  // IN: DINT
                                   INDEX := 4,  // IN: INT
                                   MLEN := 1, // IN: INT
                                   RECORD := #statDataResetParam); // INOUT: ANY

               IF NOT #statDataRecordRead.BUSY OR #statDataRecordRead.ERROR THEN
                   #statRdReq := 0;
                   #statValue := 4;
               END_IF;

           4:
               IF NOT #statRdReq AND NOT #statDataRecordRead.BUSY THEN
                   #statRdReq := 1;
               END_IF;

               #statDataRecordRead(REQ := 1,// IN: BOOL
                                   ID := #addrIn, // IN: DINT
                                   INDEX := 5, // IN: INT
                                   MLEN := 556, // IN: INT
                                   RECORD := #statDataBatteryInfo);  // INOUT: ANY

               IF NOT #statDataRecordRead.BUSY OR #statDataRecordRead.ERROR THEN
                   #statRdReq := 0;
                   IF #statDevInfoRead < 2 THEN
                       #statValue := 5;
                   ELSE
                       #statValue := 0;
                   END_IF;
               END_IF;
           5:
               IF NOT #statRdReq AND NOT #statDataRecordRead.BUSY THEN
                   #statRdReq := 1;
               END_IF;

               #statDataRecordRead(REQ := #statRdReq,  // IN: BOOL
                                   ID := #addrIn,  // IN: DINT
                                   INDEX := 6,  // IN: INT
                                   MLEN := 124, // IN: INT
                                   RECORD := #statDataDeviceInfo);  // INOUT: ANY

               IF NOT #statDataRecordRead.ERROR AND NOT #statDataRecordRead.BUSY THEN
                   #statDevInfoRead := 1;
               END_IF;

               IF NOT #statDataRecordRead.BUSY OR #statDataRecordRead.ERROR THEN
                   #statRdReq := 0;
                   #statValue := 6;
               END_IF;

           6:
               IF NOT #statRdReq AND NOT #statDataRecordRead.BUSY THEN
                   #statRdReq := 1;
               END_IF;
               #statDataRecordRead(REQ := #statRdReq,  // IN: BOOL
                                   ID := #addrIn,  // IN: DINT
                                   INDEX := 16#AFF0,  // IN: INT
                                   MLEN := 60, // IN: INT
                                   RECORD := #statDataUPSIandM);  // INOUT: ANY

               IF NOT #statDataRecordRead.ERROR AND NOT #statDataRecordRead.BUSY THEN
                   #statDevInfoRead := 1;
               END_IF;
               IF NOT #statDataRecordRead.BUSY OR #statDataRecordRead.ERROR THEN
                   #statRdReq := 0;
                   #statValue := 0;
               END_IF;
           ELSE:
               ;
       END_CASE;

       //tags datarecord index 16 write
       #HMI.State.Details.commandID := #statDataUPSCmd.commandID;
       #HMI.State.Details.parameter1 := #statDataUPSCmd.parameter1;
       #HMI.State.Details.parameter2 := #statDataUPSCmd.parameter2;

       //tags datarecord index 16#AFF0
       #HMI.State.Details.deviceHwRevision := #statDataUPSIandM.hwRevision;
       #HMI.State.Details.deviceSwRevision3 := #statDataUPSIandM.swRevision.%B0;
       #HMI.State.Details.deviceSwRevision2 := #statDataUPSIandM.swRevision.%B1;
       #HMI.State.Details.deviceSwRevision1 := #statDataUPSIandM.swRevision.%B2;
       //link data from datarecords to DB1
       //tags general (cycling datas)
       #statRetVal := DPRD_DAT(LADDR := #cyclicIOAddr, RECORD => #statCyclicData);
       IF #statRetVal <> 0 THEN
           #statStatusFLag1 := 0;
           #statStatusFLag2 := 0;
           #statDevInfoRead := 0;
           //tags datarecord index 1
           #HMI.State.bufferTime := 0;
           #HMI.State.bufferThreshold := 0;
           #HMI.State.bufferingAllowed := 0;
           //tags datarecord index 2
           //#data.batteryCapacity := 0;
           //tags datarecord index 6
           #HMI.State.maxOutCur := 0;
           //tags datarecord index 32
           #HMI.State.inputVolt := 0;
           #HMI.State.inputCur := 0;
           #HMI.State.outputVolt := 0;
           #HMI.State.loadCur := 0;
           #HMI.State.measuredChargeCur := 0;
           #HMI.State.batteryVolt := 0;
           #HMI.State.outputCur := 0;
           #HMI.State.chargeVolt := 0;
           #HMI.State.totCalcBatCap := 0;
           //#data.totCalcBatHealth := 0;
           #HMI.State.chargingOpState := 0;
           #HMI.State.endOfChargeVolt := 0;
           // Cyclic Data
           #HMI.Mode.bufferMode := 16#80;               //BZ: 4054, Solution: 16#80 to show LED off state in faceplate
           #HMI.Mode.readyForBuffering := 16#80;        //BZ: 4054 Solution: 16#80 to show LED off state in faceplate
           #HMI.State.batteryChargeLevel := 0;
       ELSE
           //tags datarecord index 1
           #HMI.State.bufferTime := #statDataBufParam.bufferTime;
           #HMI.State.bufferThreshold := INT_TO_REAL(#statDataBufParam.bufferThreshold) * 0.01;
           #HMI.State.bufferingAllowed := #statDataBufParam.bufferingAllowed;

           //tags datarecord index 2
           //HMI.State.batteryCapacity := INT_TO_REAL(#statDataBatParam.batteryCapacity) * 0.1;
           //tags datarecord index 3
           //HMI.State.chargeCur := INT_TO_REAL(#statDataChargingParam.chargeCur) * 0.001;
           //tags datarecord index 6
           #HMI.State.maxOutCur := #statDataDeviceInfo.maxOutCur;

           //tags datarecord index 32
           #HMI.State.inputVolt := INT_TO_REAL(#statDataStateInfo.inputVolt) * 0.01;
           #HMI.State.inputCur := INT_TO_REAL(#statDataStateInfo.inputCur) * 0.005;
           #HMI.State.outputVolt := INT_TO_REAL(#statDataStateInfo.outputVolt) * 0.01;
           #HMI.State.loadCur := INT_TO_REAL(#statDataStateInfo.loadCur) * 0.005;
           #HMI.State.measuredChargeCur := INT_TO_REAL(#statDataStateInfo.measuredChargeCur) * 0.001;
           #HMI.State.batteryVolt := INT_TO_REAL(#statDataStateInfo.batteryVolt) * 0.01;
           #HMI.State.outputCur := INT_TO_REAL(#statDataStateInfo.outputCur) * 0.005;
           #HMI.State.chargeVolt := INT_TO_REAL(#statDataStateInfo.chargeVolt) * 0.01;
           #HMI.State.totCalcBatCap := INT_TO_REAL(#statDataStateInfo.totalCalcBatCapacity) * 0.1;
           //#data.totCalcBatHealth := #statDataStateInfo.Reserved1;
           #HMI.State.numOfBatteries := #statDataBatteryInfo.numOfBatteries;
           #statBatteryFamily1 := DWORD_TO_BYTE(SHR(IN := #statDataBatteryInfo.batteryDetails[0].batMID, N := 24));
           #statBatteryFamily2 := DWORD_TO_BYTE(SHR(IN := #statDataBatteryInfo.batteryDetails[0].batMID, N := 16));

